REGION Network 9
   RUNG wire#powerrail
      I_Contact( "EMS".Carrier["DB401_HMI_Status".Status.CarrierStatusIndex].CommFlt )
      Contact( "EMS".Carrier["DB401_HMI_Status".Status.CarrierStatusIndex].SDC_IN.RunningREV )
      Coil( "DB401_HMI_Status".Status.RunningREV )
   END_RUNG
   // the same network as SCL:
   "DB401_HMI_Status".Status.RunningREV := NOT "EMS".Carrier["DB401_HMI_Status".Status.CarrierStatusIndex].CommFlt AND "EMS".Carrier["DB401_HMI_Status".Status.CarrierStatusIndex].SDC_IN.RunningREV;
END_REGION

REGION Network 10
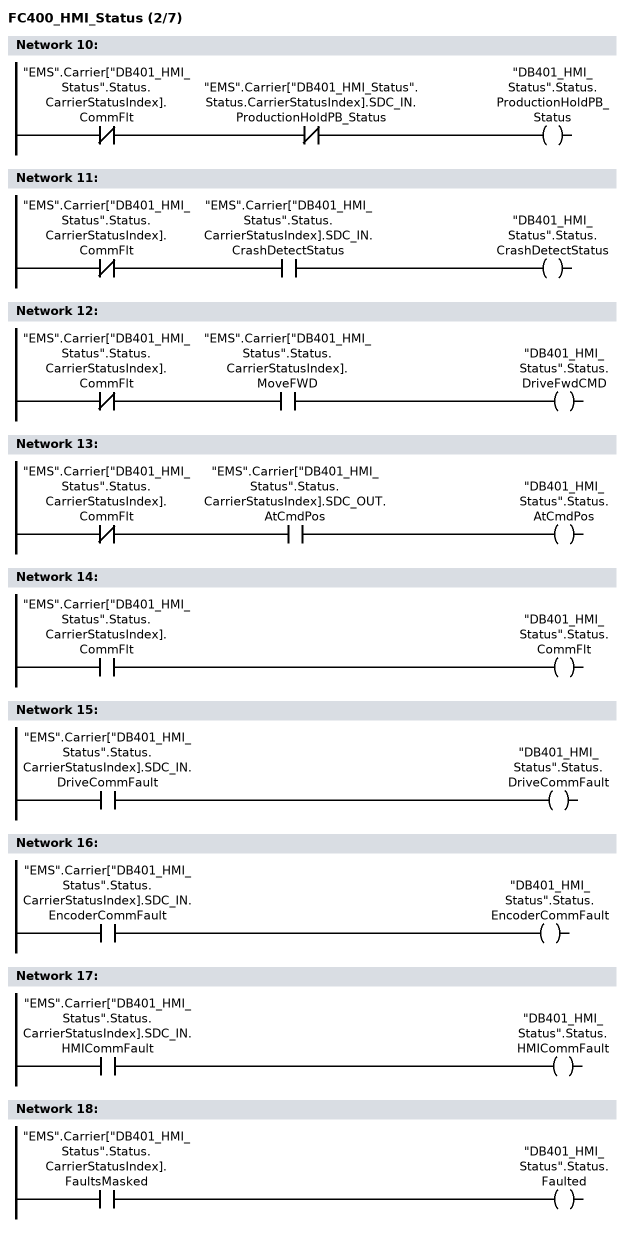
   RUNG wire#powerrail
      I_Contact( "EMS".Carrier["DB401_HMI_Status".Status.CarrierStatusIndex].CommFlt )
      I_Contact( "EMS".Carrier["DB401_HMI_Status".Status.CarrierStatusIndex].SDC_IN.ProductionHoldPB_Status )
      Coil( "DB401_HMI_Status".Status.ProductionHoldPB_Status )
   END_RUNG
   // the same network as SCL:
   "DB401_HMI_Status".Status.ProductionHoldPB_Status := NOT "EMS".Carrier["DB401_HMI_Status".Status.CarrierStatusIndex].CommFlt AND NOT "EMS".Carrier["DB401_HMI_Status".Status.CarrierStatusIndex].SDC_IN.ProductionHoldPB_Status;
END_REGION

REGION Network 11
   RUNG wire#powerrail
      I_Contact( "EMS".Carrier["DB401_HMI_Status".Status.CarrierStatusIndex].CommFlt )
      Contact( "EMS".Carrier["DB401_HMI_Status".Status.CarrierStatusIndex].SDC_IN.CrashDetectStatus )
      Coil( "DB401_HMI_Status".Status.CrashDetectStatus )
   END_RUNG
   // the same network as SCL:
   "DB401_HMI_Status".Status.CrashDetectStatus := NOT "EMS".Carrier["DB401_HMI_Status".Status.CarrierStatusIndex].CommFlt AND "EMS".Carrier["DB401_HMI_Status".Status.CarrierStatusIndex].SDC_IN.CrashDetectStatus;
END_REGION

REGION Network 12
   RUNG wire#powerrail
      I_Contact( "EMS".Carrier["DB401_HMI_Status".Status.CarrierStatusIndex].CommFlt )
      Contact( "EMS".Carrier["DB401_HMI_Status".Status.CarrierStatusIndex].MoveFWD )
      Coil( "DB401_HMI_Status".Status.DriveFwdCMD )
   END_RUNG
   // the same network as SCL:
   "DB401_HMI_Status".Status.DriveFwdCMD := NOT "EMS".Carrier["DB401_HMI_Status".Status.CarrierStatusIndex].CommFlt AND "EMS".Carrier["DB401_HMI_Status".Status.CarrierStatusIndex].MoveFWD;
END_REGION

REGION Network 13
   RUNG wire#powerrail
      I_Contact( "EMS".Carrier["DB401_HMI_Status".Status.CarrierStatusIndex].CommFlt )
      Contact( "EMS".Carrier["DB401_HMI_Status".Status.CarrierStatusIndex].SDC_OUT.AtCmdPos )
      Coil( "DB401_HMI_Status".Status.AtCmdPos )
   END_RUNG
   // the same network as SCL:
   "DB401_HMI_Status".Status.AtCmdPos := NOT "EMS".Carrier["DB401_HMI_Status".Status.CarrierStatusIndex].CommFlt AND "EMS".Carrier["DB401_HMI_Status".Status.CarrierStatusIndex].SDC_OUT.AtCmdPos;
END_REGION

REGION Network 14
   RUNG wire#powerrail
      Contact( "EMS".Carrier["DB401_HMI_Status".Status.CarrierStatusIndex].CommFlt )
      Coil( "DB401_HMI_Status".Status.CommFlt )
   END_RUNG
   // the same network as SCL:
   "DB401_HMI_Status".Status.CommFlt := "EMS".Carrier["DB401_HMI_Status".Status.CarrierStatusIndex].CommFlt;
END_REGION

REGION Network 15
   RUNG wire#powerrail
      Contact( "EMS".Carrier["DB401_HMI_Status".Status.CarrierStatusIndex].SDC_IN.DriveCommFault )
      Coil( "DB401_HMI_Status".Status.DriveCommFault )
   END_RUNG
   // the same network as SCL:
   "DB401_HMI_Status".Status.DriveCommFault := "EMS".Carrier["DB401_HMI_Status".Status.CarrierStatusIndex].SDC_IN.DriveCommFault;
END_REGION

REGION Network 16
   RUNG wire#powerrail
      Contact( "EMS".Carrier["DB401_HMI_Status".Status.CarrierStatusIndex].SDC_IN.EncoderCommFault )
      Coil( "DB401_HMI_Status".Status.EncoderCommFault )
   END_RUNG
   // the same network as SCL:
   "DB401_HMI_Status".Status.EncoderCommFault := "EMS".Carrier["DB401_HMI_Status".Status.CarrierStatusIndex].SDC_IN.EncoderCommFault;
END_REGION

REGION Network 17
   RUNG wire#powerrail
      Contact( "EMS".Carrier["DB401_HMI_Status".Status.CarrierStatusIndex].SDC_IN.HMICommFault )
      Coil( "DB401_HMI_Status".Status.HMICommFault )
   END_RUNG
   // the same network as SCL:
   "DB401_HMI_Status".Status.HMICommFault := "EMS".Carrier["DB401_HMI_Status".Status.CarrierStatusIndex].SDC_IN.HMICommFault;
END_REGION

REGION Network 18
   RUNG wire#powerrail
      Contact( "EMS".Carrier["DB401_HMI_Status".Status.CarrierStatusIndex].FaultsMasked )
      Coil( "DB401_HMI_Status".Status.Faulted )
   END_RUNG
   // the same network as SCL:
   "DB401_HMI_Status".Status.Faulted := "EMS".Carrier["DB401_HMI_Status".Status.CarrierStatusIndex].FaultsMasked;
END_REGION

REGION Network 19: PRODUCTION STOP WARNING 'H07'
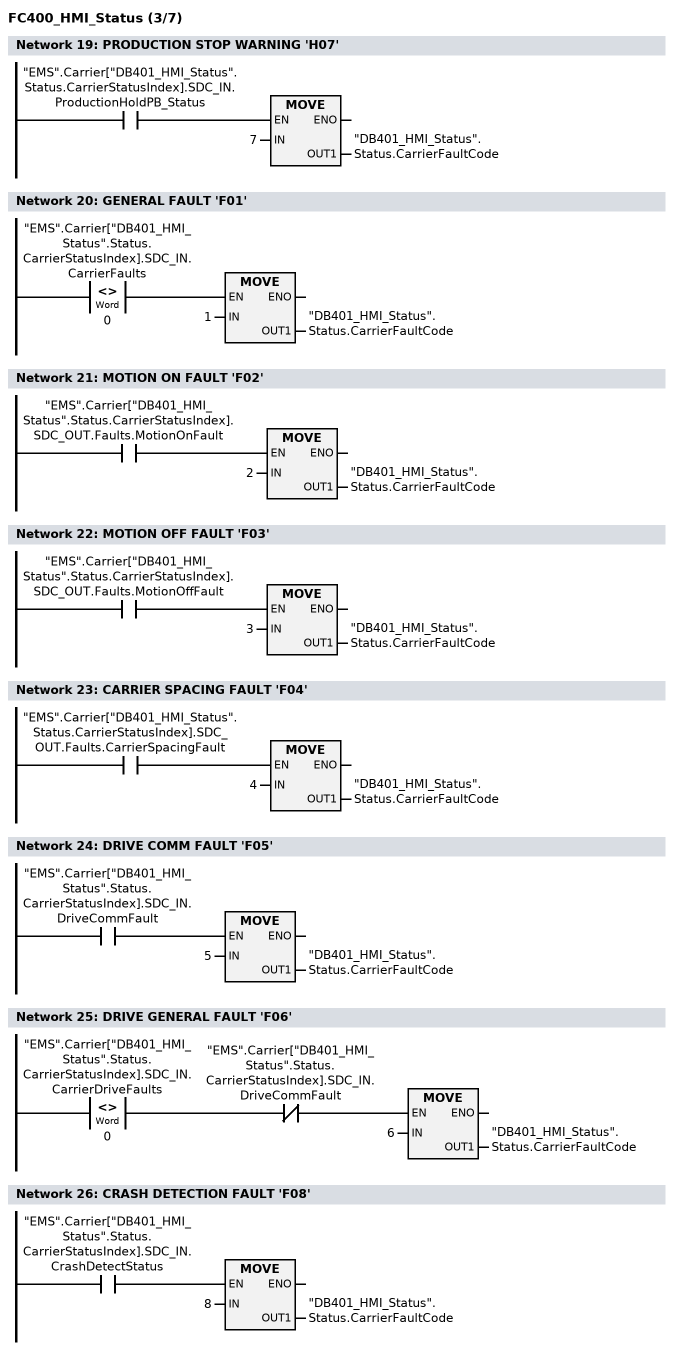
   RUNG wire#powerrail
      Contact( "EMS".Carrier["DB401_HMI_Status".Status.CarrierStatusIndex].SDC_IN.ProductionHoldPB_Status )
      Move(in := 7, out1 => "DB401_HMI_Status".Status.CarrierFaultCode)
   END_RUNG
   // the same network as SCL:
   IF "EMS".Carrier["DB401_HMI_Status".Status.CarrierStatusIndex].SDC_IN.ProductionHoldPB_Status THEN
       "DB401_HMI_Status".Status.CarrierFaultCode := 7;
   END_IF;
END_REGION

REGION Network 20: GENERAL FAULT 'F01'
   RUNG wire#powerrail
      { S7_Templates := "SrcType := Word" } NE_Contact(in1 := "EMS".Carrier["DB401_HMI_Status".Status.CarrierStatusIndex].SDC_IN.CarrierFaults, in2 := 0)
      Move(in := 1, out1 => "DB401_HMI_Status".Status.CarrierFaultCode)
   END_RUNG
   // the same network as SCL:
   IF "EMS".Carrier["DB401_HMI_Status".Status.CarrierStatusIndex].SDC_IN.CarrierFaults <> 0 THEN
       "DB401_HMI_Status".Status.CarrierFaultCode := 1;
   END_IF;
END_REGION

REGION Network 21: MOTION ON FAULT 'F02'
   RUNG wire#powerrail
      Contact( "EMS".Carrier["DB401_HMI_Status".Status.CarrierStatusIndex].SDC_OUT.Faults.MotionOnFault )
      Move(in := 2, out1 => "DB401_HMI_Status".Status.CarrierFaultCode)
   END_RUNG
   // the same network as SCL:
   IF "EMS".Carrier["DB401_HMI_Status".Status.CarrierStatusIndex].SDC_OUT.Faults.MotionOnFault THEN
       "DB401_HMI_Status".Status.CarrierFaultCode := 2;
   END_IF;
END_REGION

REGION Network 22: MOTION OFF FAULT 'F03'
   RUNG wire#powerrail
      Contact( "EMS".Carrier["DB401_HMI_Status".Status.CarrierStatusIndex].SDC_OUT.Faults.MotionOffFault )
      Move(in := 3, out1 => "DB401_HMI_Status".Status.CarrierFaultCode)
   END_RUNG
   // the same network as SCL:
   IF "EMS".Carrier["DB401_HMI_Status".Status.CarrierStatusIndex].SDC_OUT.Faults.MotionOffFault THEN
       "DB401_HMI_Status".Status.CarrierFaultCode := 3;
   END_IF;
END_REGION

REGION Network 23: CARRIER SPACING FAULT 'F04'
   RUNG wire#powerrail
      Contact( "EMS".Carrier["DB401_HMI_Status".Status.CarrierStatusIndex].SDC_OUT.Faults.CarrierSpacingFault )
      Move(in := 4, out1 => "DB401_HMI_Status".Status.CarrierFaultCode)
   END_RUNG
   // the same network as SCL:
   IF "EMS".Carrier["DB401_HMI_Status".Status.CarrierStatusIndex].SDC_OUT.Faults.CarrierSpacingFault THEN
       "DB401_HMI_Status".Status.CarrierFaultCode := 4;
   END_IF;
END_REGION

REGION Network 24: DRIVE COMM FAULT 'F05'
   RUNG wire#powerrail
      Contact( "EMS".Carrier["DB401_HMI_Status".Status.CarrierStatusIndex].SDC_IN.DriveCommFault )
      Move(in := 5, out1 => "DB401_HMI_Status".Status.CarrierFaultCode)
   END_RUNG
   // the same network as SCL:
   IF "EMS".Carrier["DB401_HMI_Status".Status.CarrierStatusIndex].SDC_IN.DriveCommFault THEN
       "DB401_HMI_Status".Status.CarrierFaultCode := 5;
   END_IF;
END_REGION

REGION Network 25: DRIVE GENERAL FAULT 'F06'
   RUNG wire#powerrail
      { S7_Templates := "SrcType := Word" } NE_Contact(in1 := "EMS".Carrier["DB401_HMI_Status".Status.CarrierStatusIndex].SDC_IN.CarrierDriveFaults, in2 := 0)
      I_Contact( "EMS".Carrier["DB401_HMI_Status".Status.CarrierStatusIndex].SDC_IN.DriveCommFault )
      Move(in := 6, out1 => "DB401_HMI_Status".Status.CarrierFaultCode)
   END_RUNG
   // the same network as SCL:
   IF ("EMS".Carrier["DB401_HMI_Status".Status.CarrierStatusIndex].SDC_IN.CarrierDriveFaults <> 0) AND NOT "EMS".Carrier["DB401_HMI_Status".Status.CarrierStatusIndex].SDC_IN.DriveCommFault THEN
       "DB401_HMI_Status".Status.CarrierFaultCode := 6;
   END_IF;
END_REGION

REGION Network 26: CRASH DETECTION FAULT 'F08'
   RUNG wire#powerrail
      Contact( "EMS".Carrier["DB401_HMI_Status".Status.CarrierStatusIndex].SDC_IN.CrashDetectStatus )
      Move(in := 8, out1 => "DB401_HMI_Status".Status.CarrierFaultCode)
   END_RUNG
   // the same network as SCL:
   IF "EMS".Carrier["DB401_HMI_Status".Status.CarrierStatusIndex].SDC_IN.CrashDetectStatus THEN
       "DB401_HMI_Status".Status.CarrierFaultCode := 8;
   END_IF;
END_REGION

REGION Network 27: DRIVE ERROR INTERNAL COMM FAULT 'F15'
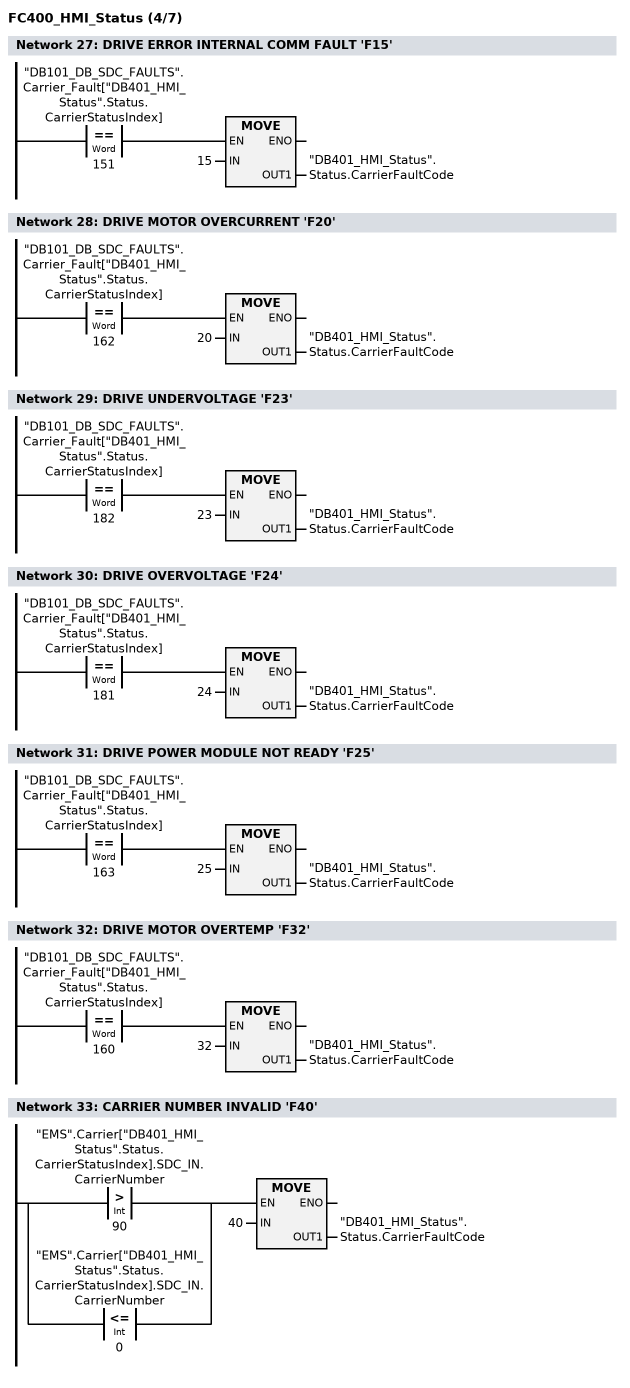
   RUNG wire#powerrail
      { S7_Templates := "SrcType := Word" } EQ_Contact(in1 := "DB101_DB_SDC_FAULTS".Carrier_Fault["DB401_HMI_Status".Status.CarrierStatusIndex], in2 := 151)
      Move(in := 15, out1 => "DB401_HMI_Status".Status.CarrierFaultCode)
   END_RUNG
   // the same network as SCL:
   IF "DB101_DB_SDC_FAULTS".Carrier_Fault["DB401_HMI_Status".Status.CarrierStatusIndex] = 151 THEN
       "DB401_HMI_Status".Status.CarrierFaultCode := 15;
   END_IF;
END_REGION

REGION Network 28: DRIVE MOTOR OVERCURRENT 'F20'
   RUNG wire#powerrail
      { S7_Templates := "SrcType := Word" } EQ_Contact(in1 := "DB101_DB_SDC_FAULTS".Carrier_Fault["DB401_HMI_Status".Status.CarrierStatusIndex], in2 := 162)
      Move(in := 20, out1 => "DB401_HMI_Status".Status.CarrierFaultCode)
   END_RUNG
   // the same network as SCL:
   IF "DB101_DB_SDC_FAULTS".Carrier_Fault["DB401_HMI_Status".Status.CarrierStatusIndex] = 162 THEN
       "DB401_HMI_Status".Status.CarrierFaultCode := 20;
   END_IF;
END_REGION

REGION Network 29: DRIVE UNDERVOLTAGE 'F23'
   RUNG wire#powerrail
      { S7_Templates := "SrcType := Word" } EQ_Contact(in1 := "DB101_DB_SDC_FAULTS".Carrier_Fault["DB401_HMI_Status".Status.CarrierStatusIndex], in2 := 182)
      Move(in := 23, out1 => "DB401_HMI_Status".Status.CarrierFaultCode)
   END_RUNG
   // the same network as SCL:
   IF "DB101_DB_SDC_FAULTS".Carrier_Fault["DB401_HMI_Status".Status.CarrierStatusIndex] = 182 THEN
       "DB401_HMI_Status".Status.CarrierFaultCode := 23;
   END_IF;
END_REGION

REGION Network 30: DRIVE OVERVOLTAGE 'F24'
   RUNG wire#powerrail
      { S7_Templates := "SrcType := Word" } EQ_Contact(in1 := "DB101_DB_SDC_FAULTS".Carrier_Fault["DB401_HMI_Status".Status.CarrierStatusIndex], in2 := 181)
      Move(in := 24, out1 => "DB401_HMI_Status".Status.CarrierFaultCode)
   END_RUNG
   // the same network as SCL:
   IF "DB101_DB_SDC_FAULTS".Carrier_Fault["DB401_HMI_Status".Status.CarrierStatusIndex] = 181 THEN
       "DB401_HMI_Status".Status.CarrierFaultCode := 24;
   END_IF;
END_REGION

REGION Network 31: DRIVE POWER MODULE NOT READY 'F25'
   RUNG wire#powerrail
      { S7_Templates := "SrcType := Word" } EQ_Contact(in1 := "DB101_DB_SDC_FAULTS".Carrier_Fault["DB401_HMI_Status".Status.CarrierStatusIndex], in2 := 163)
      Move(in := 25, out1 => "DB401_HMI_Status".Status.CarrierFaultCode)
   END_RUNG
   // the same network as SCL:
   IF "DB101_DB_SDC_FAULTS".Carrier_Fault["DB401_HMI_Status".Status.CarrierStatusIndex] = 163 THEN
       "DB401_HMI_Status".Status.CarrierFaultCode := 25;
   END_IF;
END_REGION

REGION Network 32: DRIVE MOTOR OVERTEMP 'F32'
   RUNG wire#powerrail
      { S7_Templates := "SrcType := Word" } EQ_Contact(in1 := "DB101_DB_SDC_FAULTS".Carrier_Fault["DB401_HMI_Status".Status.CarrierStatusIndex], in2 := 160)
      Move(in := 32, out1 => "DB401_HMI_Status".Status.CarrierFaultCode)
   END_RUNG
   // the same network as SCL:
   IF "DB101_DB_SDC_FAULTS".Carrier_Fault["DB401_HMI_Status".Status.CarrierStatusIndex] = 160 THEN
       "DB401_HMI_Status".Status.CarrierFaultCode := 32;
   END_IF;
END_REGION

REGION Network 33: CARRIER NUMBER INVALID 'F40'
   RUNG wire#powerrail
      { S7_Templates := "SrcType := Int" } GT_Contact(in1 := "EMS".Carrier["DB401_HMI_Status".Status.CarrierStatusIndex].SDC_IN.CarrierNumber, in2 := 90)
      wire#w1
      Move(in := 40, out1 => "DB401_HMI_Status".Status.CarrierFaultCode)
   END_RUNG
   RUNG wire#powerrail
      { S7_Templates := "SrcType := Int" } LE_Contact(in1 := "EMS".Carrier["DB401_HMI_Status".Status.CarrierStatusIndex].SDC_IN.CarrierNumber, in2 := 0)
   END_RUNG wire#w1
   // the same network as SCL:
   IF ("EMS".Carrier["DB401_HMI_Status".Status.CarrierStatusIndex].SDC_IN.CarrierNumber > 90) OR ("EMS".Carrier["DB401_HMI_Status".Status.CarrierStatusIndex].SDC_IN.CarrierNumber <= 0) THEN
       "DB401_HMI_Status".Status.CarrierFaultCode := 40;
   END_IF;
END_REGION

REGION Network 34: ENCODER FAULT 'F60'
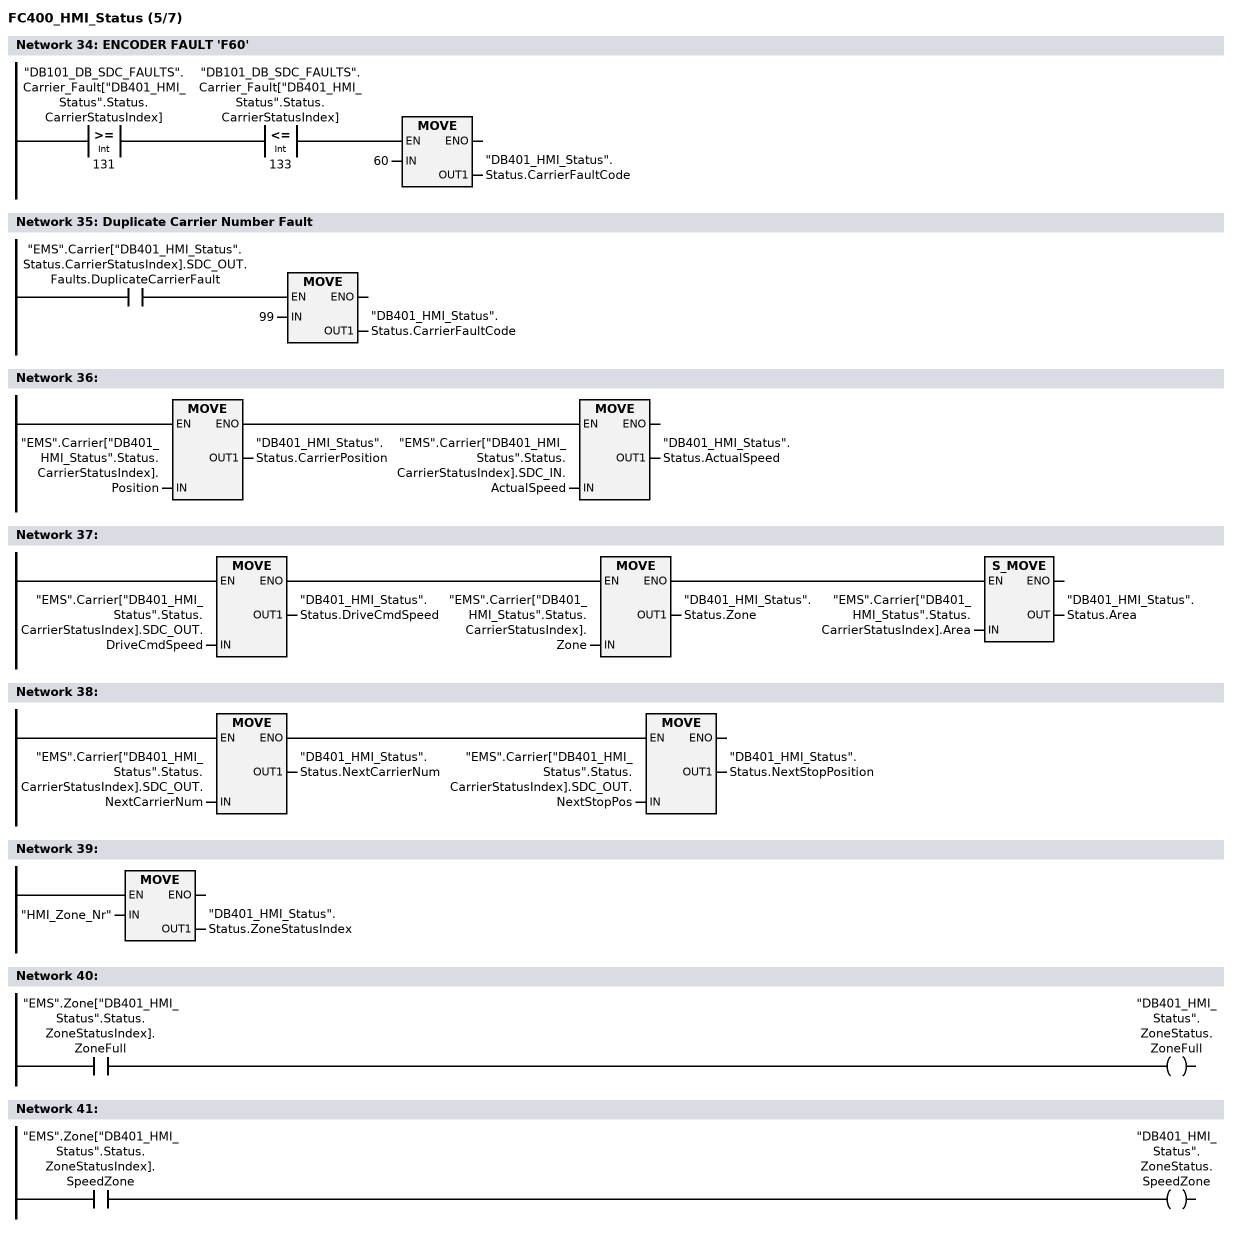
   RUNG wire#powerrail
      { S7_Templates := "SrcType := Int" } GE_Contact(in1 := "DB101_DB_SDC_FAULTS".Carrier_Fault["DB401_HMI_Status".Status.CarrierStatusIndex], in2 := 131)
      { S7_Templates := "SrcType := Int" } LE_Contact(in1 := "DB101_DB_SDC_FAULTS".Carrier_Fault["DB401_HMI_Status".Status.CarrierStatusIndex], in2 := 133)
      Move(in := 60, out1 => "DB401_HMI_Status".Status.CarrierFaultCode)
   END_RUNG
   // the same network as SCL:
   IF ("DB101_DB_SDC_FAULTS".Carrier_Fault["DB401_HMI_Status".Status.CarrierStatusIndex] >= 131) AND ("DB101_DB_SDC_FAULTS".Carrier_Fault["DB401_HMI_Status".Status.CarrierStatusIndex] <= 133) THEN
       "DB401_HMI_Status".Status.CarrierFaultCode := 60;
   END_IF;
END_REGION

REGION Network 35: Duplicate Carrier Number Fault
   RUNG wire#powerrail
      Contact( "EMS".Carrier["DB401_HMI_Status".Status.CarrierStatusIndex].SDC_OUT.Faults.DuplicateCarrierFault )
      Move(in := 99, out1 => "DB401_HMI_Status".Status.CarrierFaultCode)
   END_RUNG
   // the same network as SCL:
   IF "EMS".Carrier["DB401_HMI_Status".Status.CarrierStatusIndex].SDC_OUT.Faults.DuplicateCarrierFault THEN
       "DB401_HMI_Status".Status.CarrierFaultCode := 99;
   END_IF;
END_REGION

REGION Network 36
   RUNG wire#powerrail
      Move(in := "EMS".Carrier["DB401_HMI_Status".Status.CarrierStatusIndex].Position, out1 => "DB401_HMI_Status".Status.CarrierPosition)
      Move(in := "EMS".Carrier["DB401_HMI_Status".Status.CarrierStatusIndex].SDC_IN.ActualSpeed, out1 => "DB401_HMI_Status".Status.ActualSpeed)
   END_RUNG
   // the same network as SCL:
   "DB401_HMI_Status".Status.CarrierPosition := "EMS".Carrier["DB401_HMI_Status".Status.CarrierStatusIndex].Position;
   "DB401_HMI_Status".Status.ActualSpeed := "EMS".Carrier["DB401_HMI_Status".Status.CarrierStatusIndex].SDC_IN.ActualSpeed;
END_REGION

REGION Network 37
   RUNG wire#powerrail
      Move(in := "EMS".Carrier["DB401_HMI_Status".Status.CarrierStatusIndex].SDC_OUT.DriveCmdSpeed, out1 => "DB401_HMI_Status".Status.DriveCmdSpeed)
      Move(in := "EMS".Carrier["DB401_HMI_Status".Status.CarrierStatusIndex].Zone, out1 => "DB401_HMI_Status".Status.Zone)
      S_Move(in := "EMS".Carrier["DB401_HMI_Status".Status.CarrierStatusIndex].Area, out => "DB401_HMI_Status".Status.Area)
   END_RUNG
   // the same network as SCL:
   "DB401_HMI_Status".Status.DriveCmdSpeed := "EMS".Carrier["DB401_HMI_Status".Status.CarrierStatusIndex].SDC_OUT.DriveCmdSpeed;
   "DB401_HMI_Status".Status.Zone := "EMS".Carrier["DB401_HMI_Status".Status.CarrierStatusIndex].Zone;
   "DB401_HMI_Status".Status.Area := "EMS".Carrier["DB401_HMI_Status".Status.CarrierStatusIndex].Area;
END_REGION

REGION Network 38
   RUNG wire#powerrail
      Move(in := "EMS".Carrier["DB401_HMI_Status".Status.CarrierStatusIndex].SDC_OUT.NextCarrierNum, out1 => "DB401_HMI_Status".Status.NextCarrierNum)
      Move(in := "EMS".Carrier["DB401_HMI_Status".Status.CarrierStatusIndex].SDC_OUT.NextStopPos, out1 => "DB401_HMI_Status".Status.NextStopPosition)
   END_RUNG
   // the same network as SCL:
   "DB401_HMI_Status".Status.NextCarrierNum := "EMS".Carrier["DB401_HMI_Status".Status.CarrierStatusIndex].SDC_OUT.NextCarrierNum;
   "DB401_HMI_Status".Status.NextStopPosition := "EMS".Carrier["DB401_HMI_Status".Status.CarrierStatusIndex].SDC_OUT.NextStopPos;
END_REGION

REGION Network 39
   RUNG wire#powerrail
      Move(in := "HMI_Zone_Nr", out1 => "DB401_HMI_Status".Status.ZoneStatusIndex)
   END_RUNG
   // the same network as SCL:
   "DB401_HMI_Status".Status.ZoneStatusIndex := "HMI_Zone_Nr";
END_REGION

REGION Network 40
   RUNG wire#powerrail
      Contact( "EMS".Zone["DB401_HMI_Status".Status.ZoneStatusIndex].ZoneFull )
      Coil( "DB401_HMI_Status".ZoneStatus.ZoneFull )
   END_RUNG
   // the same network as SCL:
   "DB401_HMI_Status".ZoneStatus.ZoneFull := "EMS".Zone["DB401_HMI_Status".Status.ZoneStatusIndex].ZoneFull;
END_REGION

REGION Network 41
   RUNG wire#powerrail
      Contact( "EMS".Zone["DB401_HMI_Status".Status.ZoneStatusIndex].SpeedZone )
      Coil( "DB401_HMI_Status".ZoneStatus.SpeedZone )
   END_RUNG
   // the same network as SCL:
   "DB401_HMI_Status".ZoneStatus.SpeedZone := "EMS".Zone["DB401_HMI_Status".Status.ZoneStatusIndex].SpeedZone;
END_REGION

REGION Network 42
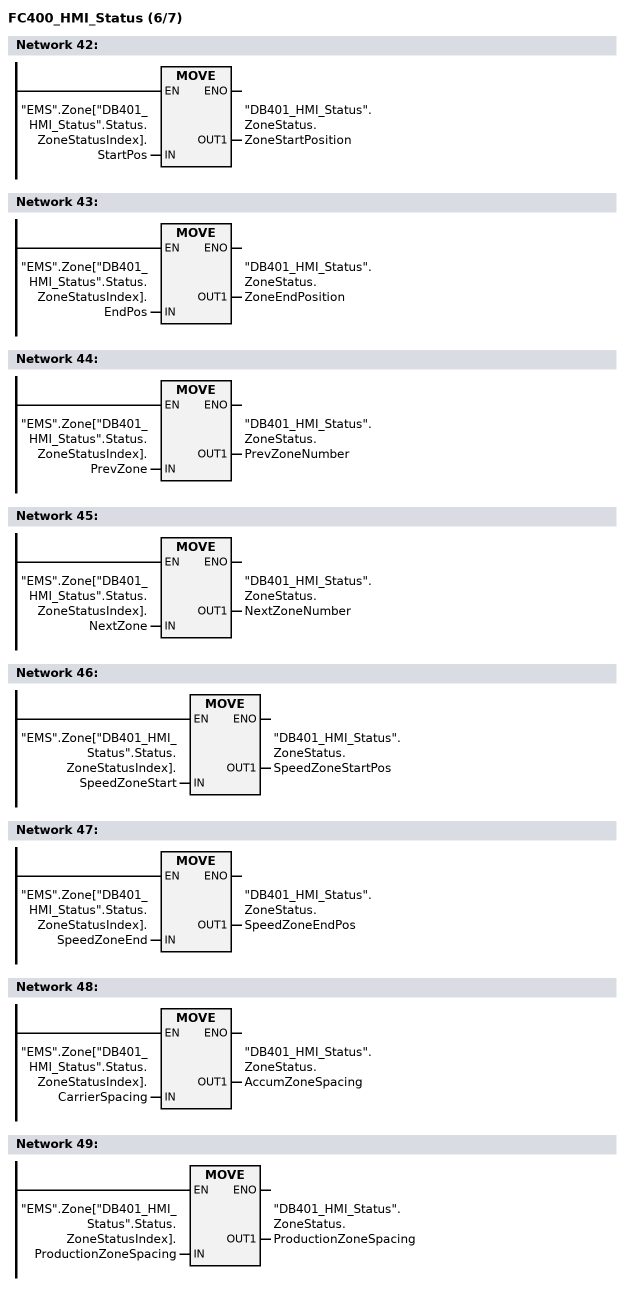
   RUNG wire#powerrail
      Move(in := "EMS".Zone["DB401_HMI_Status".Status.ZoneStatusIndex].StartPos, out1 => "DB401_HMI_Status".ZoneStatus.ZoneStartPosition)
   END_RUNG
   // the same network as SCL:
   "DB401_HMI_Status".ZoneStatus.ZoneStartPosition := "EMS".Zone["DB401_HMI_Status".Status.ZoneStatusIndex].StartPos;
END_REGION

REGION Network 43
   RUNG wire#powerrail
      Move(in := "EMS".Zone["DB401_HMI_Status".Status.ZoneStatusIndex].EndPos, out1 => "DB401_HMI_Status".ZoneStatus.ZoneEndPosition)
   END_RUNG
   // the same network as SCL:
   "DB401_HMI_Status".ZoneStatus.ZoneEndPosition := "EMS".Zone["DB401_HMI_Status".Status.ZoneStatusIndex].EndPos;
END_REGION

REGION Network 44
   RUNG wire#powerrail
      Move(in := "EMS".Zone["DB401_HMI_Status".Status.ZoneStatusIndex].PrevZone, out1 => "DB401_HMI_Status".ZoneStatus.PrevZoneNumber)
   END_RUNG
   // the same network as SCL:
   "DB401_HMI_Status".ZoneStatus.PrevZoneNumber := "EMS".Zone["DB401_HMI_Status".Status.ZoneStatusIndex].PrevZone;
END_REGION

REGION Network 45
   RUNG wire#powerrail
      Move(in := "EMS".Zone["DB401_HMI_Status".Status.ZoneStatusIndex].NextZone, out1 => "DB401_HMI_Status".ZoneStatus.NextZoneNumber)
   END_RUNG
   // the same network as SCL:
   "DB401_HMI_Status".ZoneStatus.NextZoneNumber := "EMS".Zone["DB401_HMI_Status".Status.ZoneStatusIndex].NextZone;
END_REGION

REGION Network 46
   RUNG wire#powerrail
      Move(in := "EMS".Zone["DB401_HMI_Status".Status.ZoneStatusIndex].SpeedZoneStart, out1 => "DB401_HMI_Status".ZoneStatus.SpeedZoneStartPos)
   END_RUNG
   // the same network as SCL:
   "DB401_HMI_Status".ZoneStatus.SpeedZoneStartPos := "EMS".Zone["DB401_HMI_Status".Status.ZoneStatusIndex].SpeedZoneStart;
END_REGION

REGION Network 47
   RUNG wire#powerrail
      Move(in := "EMS".Zone["DB401_HMI_Status".Status.ZoneStatusIndex].SpeedZoneEnd, out1 => "DB401_HMI_Status".ZoneStatus.SpeedZoneEndPos)
   END_RUNG
   // the same network as SCL:
   "DB401_HMI_Status".ZoneStatus.SpeedZoneEndPos := "EMS".Zone["DB401_HMI_Status".Status.ZoneStatusIndex].SpeedZoneEnd;
END_REGION

REGION Network 48
   RUNG wire#powerrail
      Move(in := "EMS".Zone["DB401_HMI_Status".Status.ZoneStatusIndex].CarrierSpacing, out1 => "DB401_HMI_Status".ZoneStatus.AccumZoneSpacing)
   END_RUNG
   // the same network as SCL:
   "DB401_HMI_Status".ZoneStatus.AccumZoneSpacing := "EMS".Zone["DB401_HMI_Status".Status.ZoneStatusIndex].CarrierSpacing;
END_REGION

REGION Network 49
   RUNG wire#powerrail
      Move(in := "EMS".Zone["DB401_HMI_Status".Status.ZoneStatusIndex].ProductionZoneSpacing, out1 => "DB401_HMI_Status".ZoneStatus.ProductionZoneSpacing)
   END_RUNG
   // the same network as SCL:
   "DB401_HMI_Status".ZoneStatus.ProductionZoneSpacing := "EMS".Zone["DB401_HMI_Status".Status.ZoneStatusIndex].ProductionZoneSpacing;
END_REGION

REGION Network 50
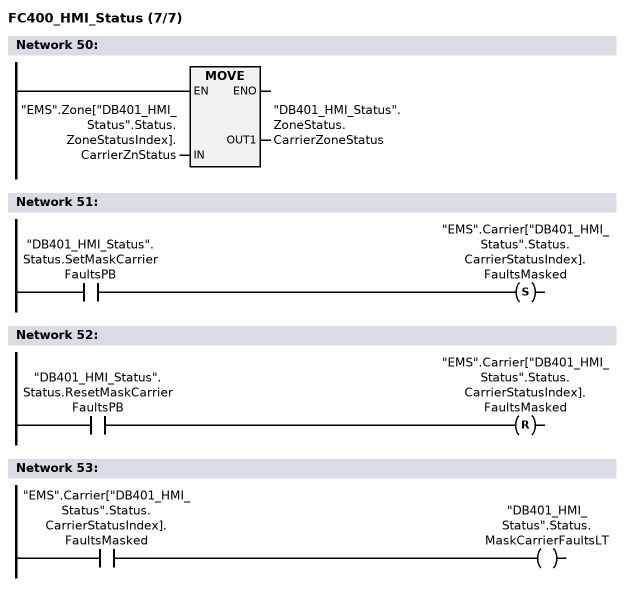
   RUNG wire#powerrail
      Move(in := "EMS".Zone["DB401_HMI_Status".Status.ZoneStatusIndex].CarrierZnStatus, out1 => "DB401_HMI_Status".ZoneStatus.CarrierZoneStatus)
   END_RUNG
   // the same network as SCL:
   "DB401_HMI_Status".ZoneStatus.CarrierZoneStatus := "EMS".Zone["DB401_HMI_Status".Status.ZoneStatusIndex].CarrierZnStatus;
END_REGION

REGION Network 51
   RUNG wire#powerrail
      Contact( "DB401_HMI_Status".Status.SetMaskCarrierFaultsPB )
      S_Coil( "EMS".Carrier["DB401_HMI_Status".Status.CarrierStatusIndex].FaultsMasked )
   END_RUNG
   // the same network as SCL:
   IF "DB401_HMI_Status".Status.SetMaskCarrierFaultsPB THEN
       "EMS".Carrier["DB401_HMI_Status".Status.CarrierStatusIndex].FaultsMasked := TRUE;
   END_IF;
END_REGION

REGION Network 52
   RUNG wire#powerrail
      Contact( "DB401_HMI_Status".Status.ResetMaskCarrierFaultsPB )
      R_Coil( "EMS".Carrier["DB401_HMI_Status".Status.CarrierStatusIndex].FaultsMasked )
   END_RUNG
   // the same network as SCL:
   IF "DB401_HMI_Status".Status.ResetMaskCarrierFaultsPB THEN
       "EMS".Carrier["DB401_HMI_Status".Status.CarrierStatusIndex].FaultsMasked := FALSE;
   END_IF;
END_REGION

REGION Network 53
   RUNG wire#powerrail
      Contact( "EMS".Carrier["DB401_HMI_Status".Status.CarrierStatusIndex].FaultsMasked )
      Coil( "DB401_HMI_Status".Status.MaskCarrierFaultsLT )
   END_RUNG
   // the same network as SCL:
   "DB401_HMI_Status".Status.MaskCarrierFaultsLT := "EMS".Carrier["DB401_HMI_Status".Status.CarrierStatusIndex].FaultsMasked;
END_REGION
END_FUNCTION

FUNCTION "FC500_FAULTS SYSTEM C1-C10" : Void   // FC500, LAD
{ S7_Optimized_Access := 'TRUE' }
VERSION : 0.1
BEGIN

REGION Network 1
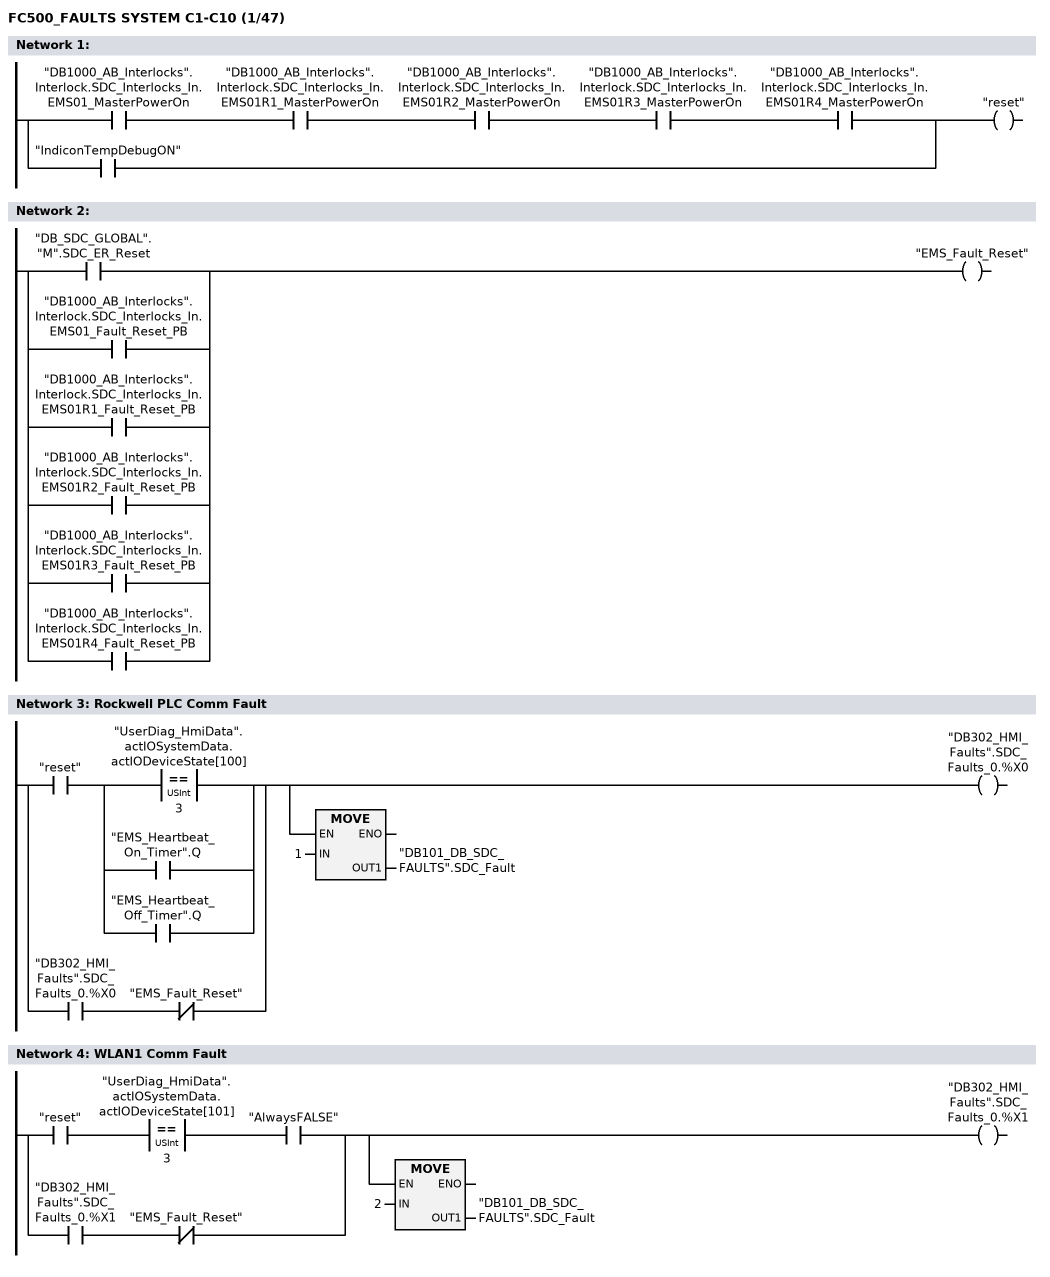
   RUNG wire#powerrail
      Contact( "DB1000_AB_Interlocks".Interlock.SDC_Interlocks_In.EMS01_MasterPowerOn )
      Contact( "DB1000_AB_Interlocks".Interlock.SDC_Interlocks_In.EMS01R1_MasterPowerOn )
      Contact( "DB1000_AB_Interlocks".Interlock.SDC_Interlocks_In.EMS01R2_MasterPowerOn )
      Contact( "DB1000_AB_Interlocks".Interlock.SDC_Interlocks_In.EMS01R3_MasterPowerOn )
      Contact( "DB1000_AB_Interlocks".Interlock.SDC_Interlocks_In.EMS01R4_MasterPowerOn )
      wire#w1
      Coil( "reset" )
   END_RUNG
   RUNG wire#powerrail
      Contact( "IndiconTempDebugON" )
   END_RUNG wire#w1
   // the same network as SCL:
   "reset" := ("DB1000_AB_Interlocks".Interlock.SDC_Interlocks_In.EMS01_MasterPowerOn AND "DB1000_AB_Interlocks".Interlock.SDC_Interlocks_In.EMS01R1_MasterPowerOn AND "DB1000_AB_Interlocks".Interlock.SDC_Interlocks_In.EMS01R2_MasterPowerOn AND "DB1000_AB_Interlocks".Interlock.SDC_Interlocks_In.EMS01R3_MasterPowerOn AND "DB1000_AB_Interlocks".Interlock.SDC_Interlocks_In.EMS01R4_MasterPowerOn) OR "IndiconTempDebugON";
END_REGION

REGION Network 2
   RUNG wire#powerrail
      Contact( "DB_SDC_GLOBAL"."M".SDC_ER_Reset )
      wire#w1
      Coil( "EMS_Fault_Reset" )
   END_RUNG
   RUNG wire#powerrail
      Contact( "DB1000_AB_Interlocks".Interlock.SDC_Interlocks_In.EMS01_Fault_Reset_PB )
   END_RUNG wire#w1
   RUNG wire#powerrail
      Contact( "DB1000_AB_Interlocks".Interlock.SDC_Interlocks_In.EMS01R1_Fault_Reset_PB )
   END_RUNG wire#w1
   RUNG wire#powerrail
      Contact( "DB1000_AB_Interlocks".Interlock.SDC_Interlocks_In.EMS01R2_Fault_Reset_PB )
   END_RUNG wire#w1
   RUNG wire#powerrail
      Contact( "DB1000_AB_Interlocks".Interlock.SDC_Interlocks_In.EMS01R3_Fault_Reset_PB )
   END_RUNG wire#w1
   RUNG wire#powerrail
      Contact( "DB1000_AB_Interlocks".Interlock.SDC_Interlocks_In.EMS01R4_Fault_Reset_PB )
   END_RUNG wire#w1
   // the same network as SCL:
   "EMS_Fault_Reset" := "DB_SDC_GLOBAL"."M".SDC_ER_Reset OR "DB1000_AB_Interlocks".Interlock.SDC_Interlocks_In.EMS01_Fault_Reset_PB OR "DB1000_AB_Interlocks".Interlock.SDC_Interlocks_In.EMS01R1_Fault_Reset_PB OR "DB1000_AB_Interlocks".Interlock.SDC_Interlocks_In.EMS01R2_Fault_Reset_PB OR "DB1000_AB_Interlocks".Interlock.SDC_Interlocks_In.EMS01R3_Fault_Reset_PB OR "DB1000_AB_Interlocks".Interlock.SDC_Interlocks_In.EMS01R4_Fault_Reset_PB;
END_REGION

REGION Network 3: Rockwell PLC Comm Fault
   RUNG wire#powerrail
      Contact( "reset" )
      wire#w1
      { S7_Templates := "SrcType := USInt" } EQ_Contact(in1 := "UserDiag_HmiData".actIOSystemData.actIODeviceState[100], in2 := 3)
      wire#w2
      Coil( "DB302_HMI_Faults".SDC_Faults_0.%X0 )
   END_RUNG
   RUNG wire#w1
      Contact( "EMS_Heartbeat_On_Timer".Q )
   END_RUNG wire#w2
   RUNG wire#w1
      Contact( "EMS_Heartbeat_Off_Timer".Q )
   END_RUNG wire#w2
   RUNG wire#powerrail
      Contact( "DB302_HMI_Faults".SDC_Faults_0.%X0 )
      I_Contact( "EMS_Fault_Reset" )
   END_RUNG wire#w2
   RUNG wire#w2
      Move(in := 1, out1 => "DB101_DB_SDC_FAULTS".SDC_Fault)
   END_RUNG
   // the same network as SCL:
   "DB302_HMI_Faults".SDC_Faults_0.%X0 := ("reset" AND (("UserDiag_HmiData".actIOSystemData.actIODeviceState[100] = 3) OR "EMS_Heartbeat_On_Timer".Q OR "EMS_Heartbeat_Off_Timer".Q)) OR ("DB302_HMI_Faults".SDC_Faults_0.%X0 AND NOT "EMS_Fault_Reset");
   IF "DB302_HMI_Faults".SDC_Faults_0.%X0 THEN "DB101_DB_SDC_FAULTS".SDC_Fault := 1; END_IF;
END_REGION

REGION Network 4: WLAN1 Comm Fault
   RUNG wire#powerrail
      Contact( "reset" )
      { S7_Templates := "SrcType := USInt" } EQ_Contact(in1 := "UserDiag_HmiData".actIOSystemData.actIODeviceState[101], in2 := 3)
      Contact( "AlwaysFALSE" )
      wire#w1
      Coil( "DB302_HMI_Faults".SDC_Faults_0.%X1 )
   END_RUNG
   RUNG wire#powerrail
      Contact( "DB302_HMI_Faults".SDC_Faults_0.%X1 )
      I_Contact( "EMS_Fault_Reset" )
   END_RUNG wire#w1
   RUNG wire#w1
      Move(in := 2, out1 => "DB101_DB_SDC_FAULTS".SDC_Fault)
   END_RUNG
   // the same network as SCL:
   "DB302_HMI_Faults".SDC_Faults_0.%X1 := ("reset" AND ("UserDiag_HmiData".actIOSystemData.actIODeviceState[101] = 3) AND "AlwaysFALSE") OR ("DB302_HMI_Faults".SDC_Faults_0.%X1 AND NOT "EMS_Fault_Reset");
   IF "DB302_HMI_Faults".SDC_Faults_0.%X1 THEN "DB101_DB_SDC_FAULTS".SDC_Fault := 2; END_IF;
END_REGION

REGION Network 5: WLAN2 Comm Fault
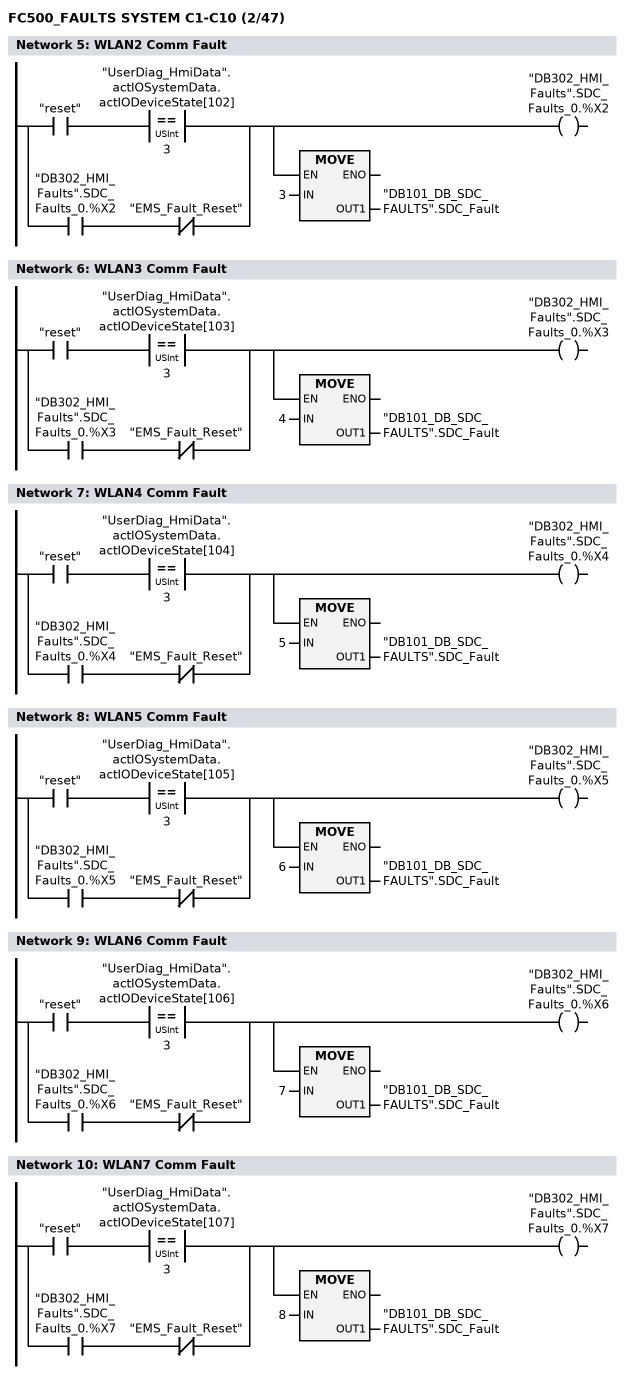
   RUNG wire#powerrail
      Contact( "reset" )
      { S7_Templates := "SrcType := USInt" } EQ_Contact(in1 := "UserDiag_HmiData".actIOSystemData.actIODeviceState[102], in2 := 3)
      wire#w1
      Coil( "DB302_HMI_Faults".SDC_Faults_0.%X2 )
   END_RUNG
   RUNG wire#powerrail
      Contact( "DB302_HMI_Faults".SDC_Faults_0.%X2 )
      I_Contact( "EMS_Fault_Reset" )
   END_RUNG wire#w1
   RUNG wire#w1
      Move(in := 3, out1 => "DB101_DB_SDC_FAULTS".SDC_Fault)
   END_RUNG
   // the same network as SCL:
   "DB302_HMI_Faults".SDC_Faults_0.%X2 := ("reset" AND ("UserDiag_HmiData".actIOSystemData.actIODeviceState[102] = 3)) OR ("DB302_HMI_Faults".SDC_Faults_0.%X2 AND NOT "EMS_Fault_Reset");
   IF "DB302_HMI_Faults".SDC_Faults_0.%X2 THEN "DB101_DB_SDC_FAULTS".SDC_Fault := 3; END_IF;
END_REGION

REGION Network 6: WLAN3 Comm Fault
   RUNG wire#powerrail
      Contact( "reset" )
      { S7_Templates := "SrcType := USInt" } EQ_Contact(in1 := "UserDiag_HmiData".actIOSystemData.actIODeviceState[103], in2 := 3)
      wire#w1
      Coil( "DB302_HMI_Faults".SDC_Faults_0.%X3 )
   END_RUNG
   RUNG wire#powerrail
      Contact( "DB302_HMI_Faults".SDC_Faults_0.%X3 )
      I_Contact( "EMS_Fault_Reset" )
   END_RUNG wire#w1
   RUNG wire#w1
      Move(in := 4, out1 => "DB101_DB_SDC_FAULTS".SDC_Fault)
   END_RUNG
   // the same network as SCL:
   "DB302_HMI_Faults".SDC_Faults_0.%X3 := ("reset" AND ("UserDiag_HmiData".actIOSystemData.actIODeviceState[103] = 3)) OR ("DB302_HMI_Faults".SDC_Faults_0.%X3 AND NOT "EMS_Fault_Reset");
   IF "DB302_HMI_Faults".SDC_Faults_0.%X3 THEN "DB101_DB_SDC_FAULTS".SDC_Fault := 4; END_IF;
END_REGION

REGION Network 7: WLAN4 Comm Fault
   RUNG wire#powerrail
      Contact( "reset" )
      { S7_Templates := "SrcType := USInt" } EQ_Contact(in1 := "UserDiag_HmiData".actIOSystemData.actIODeviceState[104], in2 := 3)
      wire#w1
      Coil( "DB302_HMI_Faults".SDC_Faults_0.%X4 )
   END_RUNG
   RUNG wire#powerrail
      Contact( "DB302_HMI_Faults".SDC_Faults_0.%X4 )
      I_Contact( "EMS_Fault_Reset" )
   END_RUNG wire#w1
   RUNG wire#w1
      Move(in := 5, out1 => "DB101_DB_SDC_FAULTS".SDC_Fault)
   END_RUNG
   // the same network as SCL:
   "DB302_HMI_Faults".SDC_Faults_0.%X4 := ("reset" AND ("UserDiag_HmiData".actIOSystemData.actIODeviceState[104] = 3)) OR ("DB302_HMI_Faults".SDC_Faults_0.%X4 AND NOT "EMS_Fault_Reset");
   IF "DB302_HMI_Faults".SDC_Faults_0.%X4 THEN "DB101_DB_SDC_FAULTS".SDC_Fault := 5; END_IF;
END_REGION
